   TextField "Text field_8" at 944,685 size 110x28; Text 'ŠKATLA 2'
   IOField "I/O field_4" at 1134,680 size 133x32; FormatPattern 999999; Unit  KOS
      ProcessValue <- "DB_STEVCI_STEVEC_SKATEL_SKATLA2"
   TextField "Text field_10" at 944,410 size 197x25; Text 'PRISOTNOST ZRAKA'
   Rectangle "Rectangle_2" at 1213,410 size 23x23
      Appearance <- "FB_Lin_FESTO_PNEVMATIKA_PRITISK_Q_izhod"
   Switch "Switch_1" at 746,167 size 165x55; CaptionText 'Switch'; TextOff 'OFF'; TextOn 'ON'
      ProcessValue <- "TimerReady"
      on Change: function_efd93a16("VARILNIK", 0, 105, 1, -1, 2)
   TextField "Text field_11" at 944,382 size 182x25; Text 'ODVIJANJE TRAKU'
   Rectangle "Rectangle_11" at 1213,382 size 23x23
      Appearance <- "NapakaOdvijanjaTrau"
   TextField "Text field_12" at 944,439 size 211x25; Text 'ČIŠČENJE ELEKTRODE'
   Rectangle "Rectangle_12" at 1213,439 size 23x23
      Appearance <- "NapakaCiscenjaElektrode"
   TextField "Text field_13" at 944,469 size 210x25; Text 'PLOŠČICA ODREZANA'
   Rectangle "Rectangle_13" at 1213,469 size 23x23
      Appearance <- "db_AKD_REZANJEPODAJANJE_PODATKI_PloscicaOdrezana"
   Button "Button_1" at 927,632 size 198x82; TextOff 'Text'
      on Click: function_efd93a16("STEVCI", 56, 120, -1, -1, 2)
   TextField "Text field_14" at 944,640 size 110x28; Text 'ŠKATLA 1'
   IOField "I/O field_5" at 1133,639 size 133x32; FormatPattern 999999; Unit  KOS
      ProcessValue <- "DB_STEVCI_STEVEC_SKATEL_SKATLA1"
   Rectangle "Rectangle_17" at 1077,643 size 23x23
      Appearance <- "FB_TekociTrak_DB_stat_skatla1Polna"
   Rectangle "Rectangle_18" at 1077,684 size 23x23
      Appearance <- "FB_TekociTrak_DB_stat_skatla2Polna"
   IOField "I/O field_9" at 297,346 size 113x44; FormatPattern 9.99; Unit s
      ProcessValue <- "FB_CYCLETIME_TimeReal"
   IOField "I/O field_8" at 297,390 size 118x23; FormatPattern 99999; Unit  KOM/H
      ProcessValue <- "FB_CYCLETIME_intfloor"
   IOField "I/O field_10" at 4,114 size 96x32; FormatPattern 1
      ProcessValue <- "Clock_5Hz"
   Group "Group" at 981,263 size 71x25
   Group "Group_1" at 981,292 size 71x25
   TextField "Text field_15" at 1073,235 size 84x25; Text 'KAMERA'
   TextField "Text field_16" at 1083,263 size 44x25; Text 'RDY'
   Rectangle "Rectangle_20" at 1133,264 size 23x23
      Appearance <- "TimerReady"
   Rectangle "Rectangle_19" at 631,361 size 135x39
      Appearance <- "FB_KAMERA_TRIG_DB_stat_CamLastValue"
   TextField "Text field_17" at 639,368 size 125x25; Text 'CAM STATUS'
   Rectangle "Rectangle_21" at 491,377 size 51x19
      Appearance <- "FB_KAMERA_TRIG_DB_io_StatusArrayCamere"
   Rectangle "Rectangle_22" at 343,531 size 17x48
      Appearance <- "FB_KAMERA_TRIG_DB_io_StatusArrayCamere"
   Polygon "Polygon_12" at 444,479 size 47x49
      Appearance <- "FB_KAMERA_TRIG_DB_io_StatusArrayCamere"
   TextField "Text field_5" at 981,263 size 44x25; Text 'RDY'
   Rectangle "Rectangle_7" at 1029,264 size 23x23
      Appearance <- "TimerReady"
   TextField "Text field_6" at 981,292 size 42x25; Text 'ERR'
   Rectangle "Rectangle_9" at 1029,293 size 23x23
      Appearance <- "WeldFault"

Template "04_PLC_StartUP" 1280x800
   Gauge "gaugeDiagStateUpdate" at 566,2 size 50x50; CaptionText 'SIMATIC'
      on Change: "CheckDiagState"()
      ProcessValue <- "@DiagnosticsIndicatorTag"
   TextField "txtTitleBar" at 16,8 size 613x32; Text 'ZAGON STROJA ... / Applikation'
   TextField "txtOperatorHeadline_1" at 768,55 size 129x23; Text 'Datum in Ura / Bediener'
   Button "btnOperator_1" at 995,56 size 40x40; TextOff '...'; PictureOff "More_Icon"
   DateTimeField "Template_Date/time field_1" at 768,72 size 208x30

screen "100_Rocno_postaja1" 1280x800, template "100_Rocno"
   TextField "Text field_1" at 729,346 size 102x25; Text 'POSTAJA1'
   Button "Button_1" at 538,135 size 200x150; TextOff 'NALAGANJE'
      on Click: SetTag("DB_HMI_ROČNI NAČIN_izbraniCilinder", 2)
   Group "Group" at 296,135 size 200x150
   Rectangle "Rectangle_4" at 678,144 size 49x30
      Appearance <- "SDAT1_oPoz2Dosezena"
   Rectangle "Rectangle_5" at 547,145 size 49x30
      Appearance <- "SDAT1_oPoz1Dosezena"
   TextField "Text field_5" at 554,147 size 30x25; Text 'B0'
   TextField "Text field_6" at 685,145 size 30x25; Text 'B1'
   Rectangle "Rectangle_6" at 548,248 size 49x30
      Appearance <- "Y2/1_NalaganjeNazanj"
   TextField "Text field_7" at 548,252 size 49x22; Text 'Y2/1'
   Rectangle "Rectangle_10" at 678,248 size 49x30
      Appearance <- "Y2/1_NalaganjeNaprej"
   TextField "Text field_11" at 679,253 size 49x22; Text 'Y2/1'
   Circle "Circle_2" at 858,253 size 24x24
      Appearance <- "PozKontaktNaKoncuLetve"
   Button "Button_3" at 770,135 size 200x150; TextOff 'PRIJEMALO'
      on Click: SetTag("DB_HMI_ROČNI NAČIN_izbraniCilinder", 3)
   Rectangle "Rectangle_7" at 911,144 size 49x30
      Appearance <- "PrijemaloKontaktaOdprto"
   Rectangle "Rectangle_8" at 780,145 size 49x30
      Appearance <- "PrijemaloKontaktaZaprto"
   TextField "Text field_8" at 787,147 size 30x25; Text 'B0'
   TextField "Text field_9" at 918,145 size 30x25; Text 'B1'
   Rectangle "Rectangle_9" at 781,248 size 49x30
      Appearance <- "Y3/1_PrijemaloKontaktaOdpri"
   TextField "Text field_10" at 781,252 size 49x22; Text 'Y3/1'
   Circle "Circle_1" at 625,253 size 24x24
      Appearance <- "PozKontaktNaKoncuLetve"
   Button "Button_2" at 296,135 size 200x150; TextOff 'ZAPORA'
      on Click: SetTag("DB_HMI_ROČNI NAČIN_izbraniCilinder", 1)
   Rectangle "Rectangle_1" at 437,144 size 49x30
      Appearance <- "ZaporaIzdelka"
   Rectangle "Rectangle_2" at 306,145 size 49x30
      Appearance <- "SprositevZaporeIzdelka"
   TextField "Text field_2" at 313,147 size 30x25; Text 'B0'
   TextField "Text field_3" at 444,145 size 30x25; Text 'B1'
   Rectangle "Rectangle_3" at 307,248 size 49x30
      Appearance <- "1Y1_OdklepZapore"
   TextField "Text field_4" at 307,252 size 49x22; Text 'Y1/1'

Template "100_Rocno" 1280x800
   TextField "txtNextBackup1" at 16,120 size 232x24; Text 'POSTAJA 1 / Option 1'
   TextField "txtNextBackup2" at 16,228 size 232x24; Text 'POSTAJA 2 / Option 1'
   TextField "txtNextBackup3" at 16,336 size 232x24; Text 'POSTAJA 3 / Option 1'
   TextField "txtNextBackup4" at 16,443 size 232x24; Text 'POSTAJA 4 / Option 1'
   IOField "ioTargetPath4" at 16,475 size 236x24; FormatPattern ??????????????????????????????????????????????????
   TextField "txtNextBackup5" at 16,551 size 232x24; Text 'Option 5 / Option 1'
   IOField "ioTargetPath5" at 16,583 size 236x24; FormatPattern ??????????????????????????????????????????????????
   TextField "txtNextBackup6" at 16,659 size 232x24; Text 'NASTAVITVE / Option 1'
   Button "btnSubNavigation1" at 2,104 size 264x109; TextOff 'Text'
      on Click: SetTag("ThirdLevelNavigationState", 1); ActivateScreen("100_Rocno_postaja1", 0)
   Button "btnSubNavigation2" at 2,211 size 264x109; TextOff 'Text'
      on Click: SetTag("ThirdLevelNavigationState", 2); ActivateScreen("102_Rocno_postaja2", 0)
   Button "btnSubNavigation3" at 1,321 size 264x109; TextOff 'Text'
      on Click: SetTag("ThirdLevelNavigationState", 3); ActivateScreen("103_Rocno_postaja3", 0)
   Button "btnSubNavigation4" at 0,432 size 264x109; TextOff 'Text'
      on Click: SetTag("ThirdLevelNavigationState", 4)
   Button "btnSubNavigation5" at 0,536 size 264x109; TextOff 'Text'
      on Click: SetTag("ThirdLevelNavigationState", 5)
   Button "btnSubNavigation6" at 2,644 size 264x109; TextOff 'Text'
      on Click: SetTag("ThirdLevelNavigationState", 6); ActivateScreen("106_Rocno_postaja6", 0)
   Gauge "gaugeDiagStateUpdate" at 566,2 size 50x50; CaptionText 'SIMATIC'
      on Change: "CheckDiagState"()
      ProcessValue <- "@DiagnosticsIndicatorTag"
   TextField "txtTitleBar" at 16,8 size 495x32; Text 'ETI C 25 - VARJENJE / Applikation'
   GraphicView "gfxNavigationIcon" at 1241,15 size 23x19; Picture "Hamburger_Icon"
   Button "btnNavigation" at 1224,0 size 56x48; TextOff 'Text'
      on Click: function_cf6f4242("GraphX_Slidein_Right", 1)
   Button "btnStartscreen" at 2,0 size 250x45; TextOff 'Text'
      on Click: "ActivateStartScreen"()
   TextField "txtStateHeadline" at 75,55 size 123x23; Text 'State / Status'
   TextField "txtRecipeHeadline" at 281,55 size 154x23; Text 'Current Recipe / Rezeptur'
   TextField "txtOperatorHeadline" at 527,55 size 129x23; Text 'Operator / Bediener'
   SymbolicIOField "ioState" at 75,72 size 119x30; TextOn '1'; TextOff '0'; TextList "Machine State"
      ProcessValue <- "RežimDelovanja"
   IOField "ioRecipe" at 281,72 size 158x30; FormatPattern ??????????????????????????????
      ProcessValue <- "CurrentRecipeName"
   IOField "ioOperator" at 527,72 size 126x30; FormatPattern ??????????????????
      ProcessValue <- "CurrentUserName"
   Button "btnState" at 202,56 size 40x40; TextOff '...'; PictureOff "More_Icon"
      on Click: "ShowOperatingModePopUp"()
   Button "btnRecipe" at 449,56 size 40x40; TextOff '...'; PictureOff "More_Icon"
      on Click: "ShowRecipePopUp"()
   Rectangle "rectState" at 0,48 size 56x56
      Appearance <- "CurrentMachineState"
   Rectangle "rectSystemDiagnosticsIndicator" at 1224,48 size 56x56
      Appearance <- "DiagState"
   GraphicIOField "gioDiagState" at 1236,60 size 32x32; PictureList "DiagState_3"
      ProcessValue <- "DiagState"
   Button "btnDiagState" at 1224,48 size 56x56; TextOff 'Text'
      on Click: ActivateScreen("30_Diagnostics", 0)
   Button "btnOperator" at 669,56 size 40x40; TextOff '...'; PictureOff "More_Icon"
      on Click: "ShowLoginPopUp"()
   TextField "txtOperatorHeadline_1" at 768,55 size 129x23; Text 'Date and Time / Bediener'
   Button "btnOperator_1" at 995,56 size 40x40; TextOff '...'; PictureOff "More_Icon"
   DateTimeField "Template_Date/time field_1" at 768,72 size 208x30
   Rectangle "rectSubNavigation1" at 0,104 size 264x109
      Appearance <- "ThirdLevelNavigationState"
   Rectangle "rectSubNavigation2" at 0,212 size 264x109
      Appearance <- "ThirdLevelNavigationState"
   Rectangle "rectSubNavigation4" at 0,428 size 264x109
      Appearance <- "ThirdLevelNavigationState"
   GraphicView "gfxPrevScreenIcon" at 1240,763 size 24x24; Picture "PrevScreen_Icon"
   Button "btnPreviousScreen" at 1223,752 size 56x48; TextOff 'Text'
      on Click: function_efd93a16()
   TextField "txtCurrentStateInfo" at 16,764 size 505x24; Text 'Optional Text about current state / Optionaler text mit aktuellem Status'
   Rectangle "rectSubNavigation4_1" at 0,536 size 264x109
      Appearance <- "ThirdLevelNavigationState"
   Rectangle "rectSubNavigation4_2" at 0,644 size 264x108
      Appearance <- "ThirdLevelNavigationState"
   Rectangle "rectSubNavigation3" at 0,320 size 264x109
      Appearance <- "ThirdLevelNavigationState"
   Rectangle "rectSubNavigation3_1" at 254,323 size 9x103
      Appearance <- "ThirdLevelNavigationState"
   Rectangle "rectSubNavigation3_2" at 254,217 size 9x103
      Appearance <- "ThirdLevelNavigationState"
   Rectangle "rectSubNavigation3_3" at 254,108 size 9x103
      Appearance <- "ThirdLevelNavigationState"
   Rectangle "rectSubNavigation3_4" at 252,644 size 9x103
      Appearance <- "ThirdLevelNavigationState"

Template "200_Rocno" 1280x800
   TextField "txtNextBackup1" at 16,120 size 232x24; Text 'POSTAJA 1 / Option 1'
   TextField "txtNextBackup2" at 16,228 size 232x24; Text 'POSTAJA 2 / Option 1'
   TextField "txtNextBackup3" at 16,336 size 232x24; Text 'POSTAJA 3 / Option 1'
   IOField "ioTargetPath3" at 16,368 size 236x24; FormatPattern ??????????????????????????????????????????????????
   TextField "txtNextBackup4" at 16,443 size 232x24; Text 'POSTAJA 4 / Option 1'
   IOField "ioTargetPath4" at 16,475 size 236x24; FormatPattern ??????????????????????????????????????????????????
   TextField "txtNextBackup5" at 16,551 size 232x24; Text 'Option 5 / Option 1'
   IOField "ioTargetPath5" at 16,583 size 236x24; FormatPattern ??????????????????????????????????????????????????
   TextField "txtNextBackup6" at 16,659 size 232x24; Text 'Option 6 / Option 1'
   IOField "ioTargetPath6" at 16,691 size 236x24; FormatPattern ??????????????????????????????????????????????????
   TextField "txtNextBackup1_1" at 2,187 size 232x24; Text 'Nalagane / Option 1'
   TextField "txtNextBackup1_2" at 6,255 size 232x24; Text 'Vrtenje / Option 1'
   TextField "txtNextBackup1_3" at 8,275 size 232x24; Text 'Varjenje / Option 1'
   Button "btnSubNavigation1" at 0,105 size 264x109; TextOff 'Text'
      on Click: SetTag("ThirdLevelNavigationState", 1)
   Button "btnSubNavigation2" at 0,215 size 264x109; TextOff 'Text'
      on Click: SetTag("ThirdLevelNavigationState", 2)
   Button "btnSubNavigation3" at 0,324 size 264x109; TextOff 'Text'
      on Click: SetTag("ThirdLevelNavigationState", 3)
   Button "btnSubNavigation4" at 1,430 size 264x109; TextOff 'Text'
      on Click: SetTag("ThirdLevelNavigationState", 4)
   Button "btnSubNavigation5" at 0,536 size 264x109; TextOff 'Text'
      on Click: SetTag("ThirdLevelNavigationState", 5)
   Button "btnSubNavigation6" at 0,644 size 264x109; TextOff 'Text'
      on Click: SetTag("ThirdLevelNavigationState", 6)
   Gauge "gaugeDiagStateUpdate" at 566,2 size 50x50; CaptionText 'SIMATIC'
      on Change: "CheckDiagState"()
      ProcessValue <- "@DiagnosticsIndicatorTag"
   TextField "txtTitleBar" at 16,8 size 495x32; Text 'ETI C 25 - VARJENJE / Applikation'
   GraphicView "gfxNavigationIcon" at 1241,15 size 23x19; Picture "Hamburger_Icon"
   Button "btnNavigation" at 1224,0 size 56x48; TextOff 'Text'
      on Click: function_cf6f4242("GraphX_Slidein_Right", 1)
   Button "btnStartscreen" at 2,0 size 250x45; TextOff 'Text'
      on Click: "ActivateStartScreen"()
   TextField "txtStateHeadline" at 75,55 size 123x23; Text 'State / Status'
   TextField "txtRecipeHeadline" at 281,55 size 154x23; Text 'Current Recipe / Rezeptur'
   TextField "txtOperatorHeadline" at 527,55 size 129x23; Text 'Operator / Bediener'
   SymbolicIOField "ioState" at 75,72 size 119x30; TextOn '1'; TextOff '0'; TextList "Machine State"
      ProcessValue <- "CurrentMachineState"
   IOField "ioRecipe" at 281,72 size 158x30; FormatPattern ??????????????????????????????
      ProcessValue <- "CurrentRecipeName"
   IOField "ioOperator" at 527,72 size 126x30; FormatPattern ??????????????????
      ProcessValue <- "CurrentUserName"
   Button "btnState" at 202,56 size 40x40; TextOff '...'; PictureOff "More_Icon"
      on Click: "ShowOperatingModePopUp"()
   Button "btnRecipe" at 449,56 size 40x40; TextOff '...'; PictureOff "More_Icon"
      on Click: "ShowRecipePopUp"()
   Rectangle "rectState" at 0,48 size 56x56
      Appearance <- "CurrentMachineState"
   Rectangle "rectSystemDiagnosticsIndicator" at 1224,48 size 56x56
      Appearance <- "DiagState"
   GraphicIOField "gioDiagState" at 1236,60 size 32x32; PictureList "DiagState_3"
      ProcessValue <- "DiagState"
   Button "btnDiagState" at 1224,48 size 56x56; TextOff 'Text'
      on Click: ActivateScreen("30_Diagnostics", 0)
   Button "btnOperator" at 669,56 size 40x40; TextOff '...'; PictureOff "More_Icon"
      on Click: "ShowLoginPopUp"()
   TextField "txtOperatorHeadline_1" at 768,55 size 129x23; Text 'Date and Time / Bediener'
   Button "btnOperator_1" at 995,56 size 40x40; TextOff '...'; PictureOff "More_Icon"
   DateTimeField "Template_Date/time field_1" at 768,72 size 208x30
   Rectangle "rectSubNavigation1" at 0,104 size 264x109
      Appearance <- "ThirdLevelNavigationState"
   Rectangle "rectSubNavigation2" at 0,212 size 264x109
      Appearance <- "ThirdLevelNavigationState"
   Rectangle "rectSubNavigation3" at 0,320 size 264x109
      Appearance <- "ThirdLevelNavigationState"
   Rectangle "rectSubNavigation4" at 0,428 size 264x109
      Appearance <- "ThirdLevelNavigationState"
   GraphicView "gfxPrevScreenIcon" at 1240,763 size 24x24; Picture "PrevScreen_Icon"
   Button "btnPreviousScreen" at 1224,751 size 56x48; TextOff 'Text'
      on Click: function_efd93a16()
   TextField "txtCurrentStateInfo" at 16,764 size 505x24; Text 'Optional Text about current state / Optionaler text mit aktuellem Status'
   Rectangle "rectSubNavigation4_1" at 0,536 size 264x109
      Appearance <- "ThirdLevelNavigationState"
   Rectangle "rectSubNavigation4_2" at 0,644 size 264x108
      Appearance <- "ThirdLevelNavigationState"

screen "102_Rocno_postaja2" 1280x800, template "100_Rocno"
   Button "Button_2" at 514,135 size 200x150; TextOff 'PODAJANJE PLOŠČICE'
      on Click: SetTag("DB_HMI_ROČNI NAČIN_izbraniCilinder", 5)
   Rectangle "Rectangle_1" at 655,144 size 49x30
      Appearance <- "ZaporaIzdelka"
   Rectangle "Rectangle_2" at 524,145 size 49x30
      Appearance <- "SprositevZaporeIzdelka"
   TextField "Text field_2" at 531,147 size 30x25; Text 'B0'
   TextField "Text field_3" at 662,145 size 30x25; Text 'B1'
   Rectangle "Rectangle_3" at 525,248 size 49x30
      Appearance <- "Y2/1_dovajanjeKontaktovNazaj"
   TextField "Text field_4" at 525,252 size 49x22; Text 'Y1/2'
   Rectangle "Rectangle_14" at 655,248 size 49x30
      Appearance <- "Y2_1_dovajanjeKntaktovNaprej"
   TextField "Text field_15" at 655,252 size 49x22; Text 'Y1/2'
   Button "Button_10" at 732,135 size 200x150; TextOff 'PODAJANJE/REZANJE TRAKA'
      on Click: SetTag("DB_HMI_ROČNI NAČIN_izbraniCilinder", 22)
   Button "Button_1" at 299,135 size 200x150; TextOff 'ČIŠČENJE ELEKTRODE'
      on Click: SetTag("DB_HMI_ROČNI NAČIN_izbraniCilinder", 220)
   Rectangle "Rectangle_4" at 309,145 size 49x30
      Appearance <- "SenzorOdvijanjaCiscenjeElektrode"
   TextField "Text field_5" at 316,147 size 30x25; Text 'B0'
   TextField "Text field_1" at 742,250 size 21x25; Text 'M'
   Rectangle "Rectangle_5" at 740,141 size 38x28
      Appearance <- "FB_STARTUP_DB_DeviceState_mySTATE{5}"
   TextField "Text field_6" at 744,145 size 29x22; Text 'PN'
   Rectangle "Rectangle_29" at 789,141 size 38x28
      Appearance <- "FB_AKD_REZANJEPODAJANJE_iAKD_PODATKI_TO_SIEMENS_HomePosSet"
   TextField "Text field_29" at 800,145 size 17x22; Text 'H'
   Rectangle "Rectangle_33" at 880,141 size 38x28
      Appearance <- "FB_AKD_REZANJEPODAJANJE_iAKD_PODATKI_TO_SIEMENS_WarningPreent"
   TextField "Text field_33" at 888,144 size 21x22; Text 'W'
   Rectangle "Rectangle_30" at 835,141 size 38x28
      Appearance <- "FB_AKD_DB_RezanjePodajanje_iAKD_PODATKI_TO_SIEMENS_FaultPresent"
   TextField "Text field_30" at 835,145 size 39x22; Text 'ERR'

screen "103_Rocno_postaja3" 1280x800, template "100_Rocno"
   Button "Button_2" at 296,135 size 200x150; TextOff 'DVIG/SPUST ELEKTRODE'
      on Click: SetTag("DB_HMI_ROČNI NAČIN_izbraniCilinder", 6)
   Rectangle "Rectangle_1" at 437,144 size 49x30
      Appearance <- "FB_KEYENCE_GT2_ODMIKVARJENJA_oPoz3Dosezena"
   Rectangle "Rectangle_2" at 306,145 size 49x30
      Appearance <- "FB_KEYENCE_GT2_ODMIKVARJENJA_oPoz1Dosezena"
   TextField "Text field_2" at 313,147 size 30x25; Text 'B0'
   TextField "Text field_3" at 444,145 size 30x25; Text 'B1'
   Rectangle "Rectangle_3" at 307,248 size 49x30
      Appearance <- "Y1/3_odmičniCilinderVarjenje_GOR"
   TextField "Text field_4" at 307,252 size 49x22; Text 'Y1/3'
   Rectangle "Rectangle_14" at 437,248 size 49x30
      Appearance <- "Y1/3_odmičniCilinderVarjenjeDOL"
   TextField "Text field_15" at 437,252 size 49x22; Text 'Y1/3'
   Button "Button_1" at 537,135 size 200x150; TextOff 'PORAVNANA KONTAKTA'
      on Click: SetTag("DB_HMI_ROČNI NAČIN_izbraniCilinder", 7)
   Rectangle "Rectangle_4" at 678,144 size 49x30
      Appearance <- "PozKontaktNaprej"
   Rectangle "Rectangle_5" at 547,145 size 49x30
      Appearance <- "PozKontaktNazaj"
   TextField "Text field_5" at 554,147 size 30x25; Text 'B0'
   TextField "Text field_6" at 685,145 size 30x25; Text 'B1'
   Rectangle "Rectangle_6" at 548,248 size 49x30
      Appearance <- "Y2/3_PozicioniranjeKontaktovNazaj"
   TextField "Text field_7" at 548,252 size 49x22; Text 'Y2/1'
   Rectangle "Rectangle_10" at 678,248 size 49x30
      Appearance <- "Y2/3_PozicioniranjeKontaktovNaprej"
   TextField "Text field_11" at 679,253 size 49x22; Text 'Y2/1'
   Button "Button_5" at 778,135 size 200x150; TextOff 'ODKLEP/ZAKLEP KONUSA'
      on Click: SetTag("DB_HMI_ROČNI NAČIN_izbraniCilinder", 8)
   Rectangle "Rectangle_15" at 919,144 size 49x30
      Appearance <- "FB_KEYENCE_GT2_odmikKonusaKroznika_oPoz2Dosezena"
   Rectangle "Rectangle_16" at 788,145 size 49x30
      Appearance <- "FB_KEYENCE_GT2_odmikKonusaKroznika_oPoz1Dosezena"
   TextField "Text field_16" at 795,147 size 30x25; Text 'B0'
   TextField "Text field_17" at 926,145 size 30x25; Text 'B1'
   Rectangle "Rectangle_17" at 789,248 size 49x30
      Appearance <- "Y1/3_OdmičniCilinderKonusa"
   TextField "Text field_18" at 789,252 size 49x22; Text 'Y1/3'
   Button "Button_4" at 1020,135 size 200x150; TextOff 'ODKLEP VSTAVLJANJE KONTAKTA'
      on Click: SetTag("DB_HMI_ROČNI NAČIN_izbraniCilinder", 9)
   Rectangle "Rectangle_12" at 1030,145 size 49x30
      Appearance <- "DrzanjeKontakta"
   TextField "Text field_12" at 1037,147 size 30x25; Text 'B0'
   Rectangle "Rectangle_13" at 1031,248 size 49x30
      Appearance <- "Y3/3_OdpiranjeDržalaKomada"
   TextField "Text field_14" at 1031,252 size 49x22; Text 'Y3/3'
   Button "Button_3" at 296,307 size 200x150; TextOff 'ODKLEP IZMETA KONTAKTA'
      on Click: SetTag("DB_HMI_ROČNI NAČIN_izbraniCilinder", 10)
   Rectangle "Rectangle_7" at 306,317 size 49x30
      Appearance <- "DrzanjeIzmetKontakta"
   TextField "Text field_8" at 313,319 size 30x25; Text 'B0'
   Rectangle "Rectangle_8" at 307,420 size 49x30
      Appearance <- "Y4/3_OdpiranjeIzmetaKontakta"
   TextField "Text field_9" at 307,424 size 49x22; Text 'Y4/3'
   Button "Button_6" at 537,307 size 200x150; TextOff 'ODKLEP IZMETA KONTAKTA'
      on Click: SetTag("DB_HMI_ROČNI NAČIN_izbraniCilinder", 11)
   Rectangle "Rectangle_9" at 547,317 size 49x30
      Appearance <- "IzmetKontaktaNazaj"
   TextField "Text field_10" at 554,319 size 30x25; Text 'B0'
   Rectangle "Rectangle_11" at 548,420 size 49x30
      Appearance <- "Y5/3_IzmetKomadov"
   TextField "Text field_13" at 548,424 size 49x22; Text 'Y5/3'
   Button "Button_7" at 778,307 size 200x150; TextOff 'DRČA'
      on Click: SetTag("DB_HMI_ROČNI NAČIN_izbraniCilinder", 12)
   Rectangle "Rectangle_18" at 919,316 size 49x30
      Appearance <- "DrcaDobriKosi"
   Rectangle "Rectangle_19" at 788,317 size 49x30
      Appearance <- "DrscaSLabiKosi"
   TextField "Text field_19" at 795,319 size 30x25; Text 'B0'
   TextField "Text field_20" at 926,317 size 30x25; Text 'B1'
   Rectangle "Rectangle_20" at 789,420 size 49x30
      Appearance <- "Y6/3_LoputaSlabi"
   TextField "Text field_21" at 789,424 size 49x22; Text 'Y6/3'
   Rectangle "Rectangle_21" at 919,420 size 49x30
      Appearance <- "Y6/3_LoputaDobri"
   TextField "Text field_22" at 920,425 size 49x22; Text 'Y6/3'
   Button "Button_8" at 295,539 size 200x150; TextOff 'VRTENJE MIZE'
      on Click: SetTag("DB_HMI_ROČNI NAČIN_izbraniCilinder", 20)
   Rectangle "Rectangle_22" at 300,549 size 38x28
      Appearance <- "FB_STARTUP_DB_DeviceState_mySTATE{7}"
   TextField "Text field_1" at 304,553 size 29x22; Text 'PN'
   Button "Button_9" at 537,539 size 200x150; TextOff 'VRTENJE ELEKTRODE'
      on Click: SetTag("DB_HMI_ROČNI NAČIN_izbraniCilinder", 21)
   Button "Button_10" at 778,539 size 200x150; TextOff 'PODAJANJE/REZANJE TRAKA'
      on Click: SetTag("DB_HMI_ROČNI NAČIN_izbraniCilinder", 22)
   Rectangle "Rectangle_23" at 544,551 size 38x28
      Appearance <- "FB_STARTUP_DB_DeviceState_mySTATE{8}"
   TextField "Text field_23" at 548,555 size 29x22; Text 'PN'
   Rectangle "Rectangle_24" at 787,552 size 38x28
      Appearance <- "FB_STARTUP_DB_DeviceState_mySTATE{5}"
   TextField "Text field_24" at 791,556 size 29x22; Text 'PN'
   Rectangle "Rectangle_25" at 347,549 size 38x28
      Appearance <- "FB_AKD_VrtenjeKroznika_iAKD_PODATKI_TO_SIEMENS_HomePosSet"
   TextField "Text field_25" at 358,552 size 17x22; Text 'H'
   Rectangle "Rectangle_26" at 393,549 size 38x28
      Appearance <- "FB_AKD_Kroznik_iAKD_PODATKI_TO_SIEMENS_FaultPresent"
   TextField "Text field_26" at 393,552 size 39x22; Text 'ERR'
   Rectangle "Rectangle_27" at 592,550 size 38x28
      Appearance <- "FB_AKD_VrtenjeELektrode_iAKD_PODATKI_TO_SIEMENS_HomePosSet"
   TextField "Text field_27" at 603,553 size 17x22; Text 'H'
   Rectangle "Rectangle_28" at 638,550 size 38x28
      Appearance <- "FB_AKD_DB_elektroda_iAKD_PODATKI_TO_SIEMENS_FaultPresent"
   TextField "Text field_28" at 638,553 size 39x22; Text 'ERR'
   Rectangle "Rectangle_29" at 836,552 size 38x28
      Appearance <- "FB_AKD_REZANJEPODAJANJE_iAKD_PODATKI_TO_SIEMENS_HomePosSet"
   TextField "Text field_29" at 847,555 size 17x22; Text 'H'
   Rectangle "Rectangle_30" at 882,552 size 38x28
      Appearance <- "FB_AKD_DB_RezanjePodajanje_iAKD_PODATKI_TO_SIEMENS_FaultPresent"
   TextField "Text field_30" at 882,555 size 39x22; Text 'ERR'
   Rectangle "Rectangle_31" at 441,549 size 38x28
      Appearance <- "FB_AKD_Kroznik_iAKD_PODATKI_TO_SIEMENS_WarningPreent"
   TextField "Text field_31" at 449,552 size 21x22; Text 'W'
   Rectangle "Rectangle_32" at 686,549 size 38x28
      Appearance <- "FB_AKD_VrtenjeELektrode_iAKD_PODATKI_TO_SIEMENS_WarningPreent"
   TextField "Text field_32" at 694,552 size 21x22; Text 'W'
   Rectangle "Rectangle_33" at 927,552 size 38x28
      Appearance <- "FB_AKD_REZANJEPODAJANJE_iAKD_PODATKI_TO_SIEMENS_WarningPreent"
   TextField "Text field_33" at 935,555 size 21x22; Text 'W'
   TextField "Text field_34" at 332,664 size 138x25; Text 'onemogoceno'
      Visibility <- "FB_AKD_VrtenjeKroznika_OmogociHome"
   Switch "Switch_1" at 296,694 size 198x55; CaptionText 'START HOME'; TextOff 'OFF'; TextOn 'ON'
      ProcessValue <- "DB_HMI_Kroznik_bStartHomming"
      Appearance <- "FB_AKD_VrtenjeKroznika_OmogociHome"
      Visibility <- "FB_AKD_VrtenjeKroznika_OmogociHome"

